// TIA Portal project "Canarias Skills" (V17) (continued)
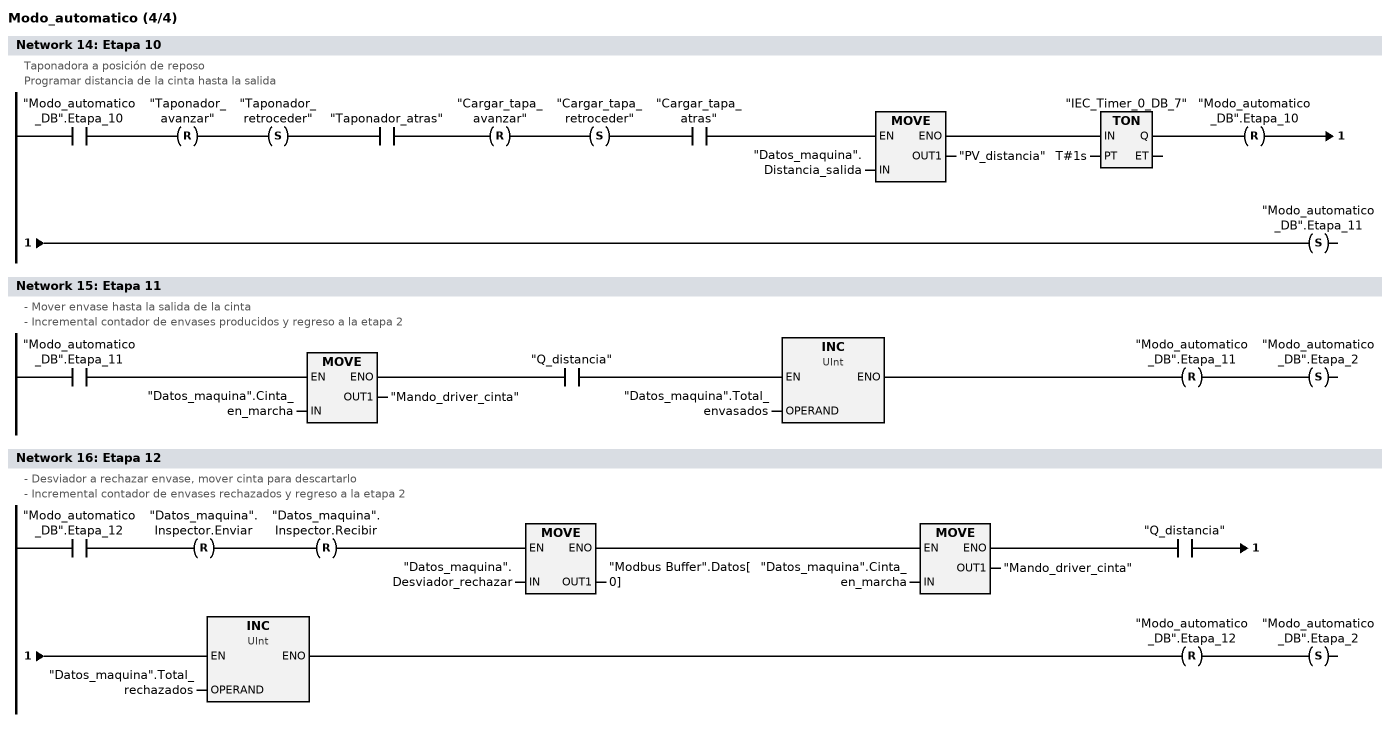
   IF "Modo_automatico_DB".Etapa_10 THEN
       "Taponador_avanzar" := FALSE;
       "Taponador_retroceder" := TRUE;
   END_IF;
   #_w1 := "Modo_automatico_DB".Etapa_10 AND "Taponador_atras";
   IF #_w1 THEN
       "Cargar_tapa_avanzar" := FALSE;
       "Cargar_tapa_retroceder" := TRUE;
   END_IF;
   #_w2 := #_w1 AND "Cargar_tapa_atras";
   IF #_w2 THEN "PV_distancia" := "Datos_maquina".Distancia_salida; END_IF;
   "IEC_Timer_0_DB_7".TON(IN := #_w2, PT := T#1s);
   IF "IEC_Timer_0_DB_7".Q THEN
       "Modo_automatico_DB".Etapa_10 := FALSE;
       "Modo_automatico_DB".Etapa_11 := TRUE;
   END_IF;
END_REGION

REGION Network 15: Etapa 11
   // - Mover envase hasta la salida de la cinta
   // - Incremental contador de envases producidos y regreso a la etapa 2
   RUNG wire#powerrail
      Contact( "Modo_automatico_DB".Etapa_11 )
      Move(in := "Datos_maquina".Cinta_en_marcha, out1 => "Mando_driver_cinta")
      Contact( "Q_distancia" )
      { S7_Templates := "DestType := UInt" } Inc( "Datos_maquina".Total_envasados )
      R_Coil( "Modo_automatico_DB".Etapa_11 )
      S_Coil( "Modo_automatico_DB".Etapa_2 )
   END_RUNG
   // the same network as SCL:
   IF "Modo_automatico_DB".Etapa_11 THEN "Mando_driver_cinta" := "Datos_maquina".Cinta_en_marcha; END_IF;
   IF "Modo_automatico_DB".Etapa_11 AND "Q_distancia" THEN
       "Datos_maquina".Total_envasados := "Datos_maquina".Total_envasados + 1;
   END_IF;
   #_w1 := "Modo_automatico_DB".Etapa_11 AND "Q_distancia";
   IF #_w1 THEN
       "Modo_automatico_DB".Etapa_11 := FALSE;
       "Modo_automatico_DB".Etapa_2 := TRUE;
   END_IF;
END_REGION

REGION Network 16: Etapa 12
   // - Desviador a rechazar envase, mover cinta para descartarlo
   // - Incremental contador de envases rechazados y regreso a la etapa 2
   RUNG wire#powerrail
      Contact( "Modo_automatico_DB".Etapa_12 )
      R_Coil( "Datos_maquina".Inspector.Enviar )
      R_Coil( "Datos_maquina".Inspector.Recibir )
      Move(in := "Datos_maquina".Desviador_rechazar, out1 => "Modbus Buffer".Datos[0])
      Move(in := "Datos_maquina".Cinta_en_marcha, out1 => "Mando_driver_cinta")
      Contact( "Q_distancia" )
      { S7_Templates := "DestType := UInt" } Inc( "Datos_maquina".Total_rechazados )
      R_Coil( "Modo_automatico_DB".Etapa_12 )
      S_Coil( "Modo_automatico_DB".Etapa_2 )
   END_RUNG
   // the same network as SCL:
   IF "Modo_automatico_DB".Etapa_12 THEN
       "Datos_maquina".Inspector.Enviar := FALSE;
       "Datos_maquina".Inspector.Recibir := FALSE;
       "Modbus Buffer".Datos[0] := "Datos_maquina".Desviador_rechazar;
       "Mando_driver_cinta" := "Datos_maquina".Cinta_en_marcha;
   END_IF;
   IF "Modo_automatico_DB".Etapa_12 AND "Q_distancia" THEN
       "Datos_maquina".Total_rechazados := "Datos_maquina".Total_rechazados + 1;
   END_IF;
   #_w1 := "Modo_automatico_DB".Etapa_12 AND "Q_distancia";
   IF #_w1 THEN
       "Modo_automatico_DB".Etapa_12 := FALSE;
       "Modo_automatico_DB".Etapa_2 := TRUE;
   END_IF;
END_REGION
END_FUNCTION_BLOCK

FUNCTION "Inicializar maquina" : Void   // FC1, LAD
{ S7_Optimized_Access := 'TRUE' }
VERSION : 0.1
BEGIN

REGION Network 1
   // Variador cinta, en servicio y detenido
   // Desviador en posición de aceptar envase
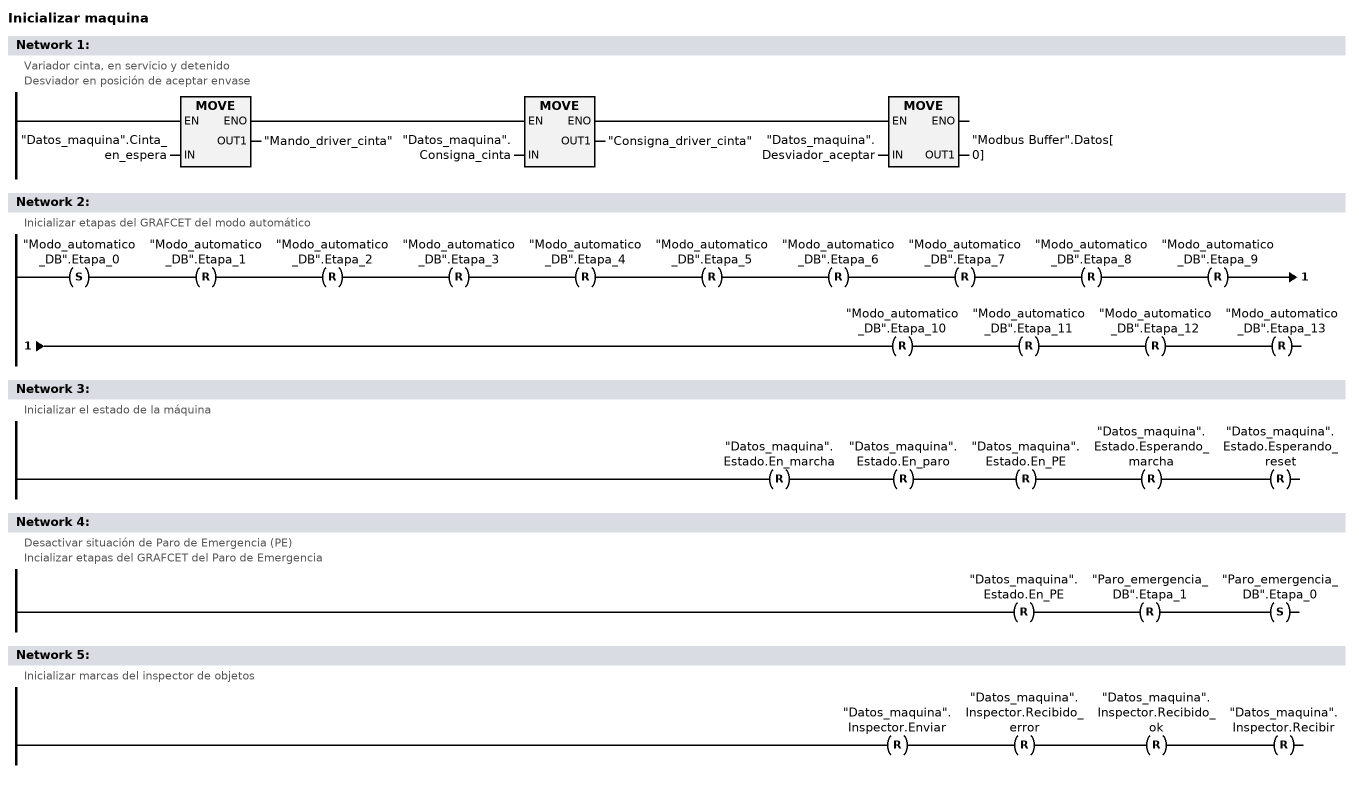
   RUNG wire#powerrail
      Move(in := "Datos_maquina".Cinta_en_espera, out1 => "Mando_driver_cinta")
      Move(in := "Datos_maquina".Consigna_cinta, out1 => "Consigna_driver_cinta")
      Move(in := "Datos_maquina".Desviador_aceptar, out1 => "Modbus Buffer".Datos[0])
   END_RUNG
   // the same network as SCL:
   "Mando_driver_cinta" := "Datos_maquina".Cinta_en_espera;
   "Consigna_driver_cinta" := "Datos_maquina".Consigna_cinta;
   "Modbus Buffer".Datos[0] := "Datos_maquina".Desviador_aceptar;
END_REGION

REGION Network 2
   // Inicializar etapas del GRAFCET del modo automático
   RUNG wire#powerrail
      S_Coil( "Modo_automatico_DB".Etapa_0 )
      R_Coil( "Modo_automatico_DB".Etapa_1 )
      R_Coil( "Modo_automatico_DB".Etapa_2 )
      R_Coil( "Modo_automatico_DB".Etapa_3 )
      R_Coil( "Modo_automatico_DB".Etapa_4 )
      R_Coil( "Modo_automatico_DB".Etapa_5 )
      R_Coil( "Modo_automatico_DB".Etapa_6 )
      R_Coil( "Modo_automatico_DB".Etapa_7 )
      R_Coil( "Modo_automatico_DB".Etapa_8 )
      R_Coil( "Modo_automatico_DB".Etapa_9 )
      R_Coil( "Modo_automatico_DB".Etapa_10 )
      R_Coil( "Modo_automatico_DB".Etapa_11 )
      R_Coil( "Modo_automatico_DB".Etapa_12 )
      R_Coil( "Modo_automatico_DB".Etapa_13 )
   END_RUNG
   // the same network as SCL:
   "Modo_automatico_DB".Etapa_0 := TRUE;
   "Modo_automatico_DB".Etapa_1 := FALSE;
   "Modo_automatico_DB".Etapa_2 := FALSE;
   "Modo_automatico_DB".Etapa_3 := FALSE;
   "Modo_automatico_DB".Etapa_4 := FALSE;
   "Modo_automatico_DB".Etapa_5 := FALSE;
   "Modo_automatico_DB".Etapa_6 := FALSE;
   "Modo_automatico_DB".Etapa_7 := FALSE;
   "Modo_automatico_DB".Etapa_8 := FALSE;
   "Modo_automatico_DB".Etapa_9 := FALSE;
   "Modo_automatico_DB".Etapa_10 := FALSE;
   "Modo_automatico_DB".Etapa_11 := FALSE;
   "Modo_automatico_DB".Etapa_12 := FALSE;
   "Modo_automatico_DB".Etapa_13 := FALSE;
END_REGION

REGION Network 3
   // Inicializar el estado de la máquina
   RUNG wire#powerrail
      R_Coil( "Datos_maquina".Estado.En_marcha )
      R_Coil( "Datos_maquina".Estado.En_paro )
      R_Coil( "Datos_maquina".Estado.En_PE )
      R_Coil( "Datos_maquina".Estado.Esperando_marcha )
      R_Coil( "Datos_maquina".Estado.Esperando_reset )
   END_RUNG
   // the same network as SCL:
   "Datos_maquina".Estado.En_marcha := FALSE;
   "Datos_maquina".Estado.En_paro := FALSE;
   "Datos_maquina".Estado.En_PE := FALSE;
   "Datos_maquina".Estado.Esperando_marcha := FALSE;
   "Datos_maquina".Estado.Esperando_reset := FALSE;
END_REGION

REGION Network 4
   // Desactivar situación de Paro de Emergencia (PE)
   // Incializar etapas del GRAFCET del Paro de Emergencia
   RUNG wire#powerrail
      R_Coil( "Datos_maquina".Estado.En_PE )
      R_Coil( "Paro_emergencia_DB".Etapa_1 )
      S_Coil( "Paro_emergencia_DB".Etapa_0 )
   END_RUNG
   // the same network as SCL:
   "Datos_maquina".Estado.En_PE := FALSE;
   "Paro_emergencia_DB".Etapa_1 := FALSE;
   "Paro_emergencia_DB".Etapa_0 := TRUE;
END_REGION

REGION Network 5
   // Inicializar marcas del inspector de objetos
   RUNG wire#powerrail
      R_Coil( "Datos_maquina".Inspector.Enviar )
      R_Coil( "Datos_maquina".Inspector.Recibido_error )
      R_Coil( "Datos_maquina".Inspector.Recibido_ok )
      R_Coil( "Datos_maquina".Inspector.Recibir )
   END_RUNG
   // the same network as SCL:
   "Datos_maquina".Inspector.Enviar := FALSE;
   "Datos_maquina".Inspector.Recibido_error := FALSE;
   "Datos_maquina".Inspector.Recibido_ok := FALSE;
   "Datos_maquina".Inspector.Recibir := FALSE;
END_REGION
END_FUNCTION

FUNCTION "Modo manual" : Void   // FC2, LAD
{ S7_Optimized_Access := 'TRUE' }
VERSION : 0.1
BEGIN

REGION Network 1: Maniobra manual de la neumática desde HMI
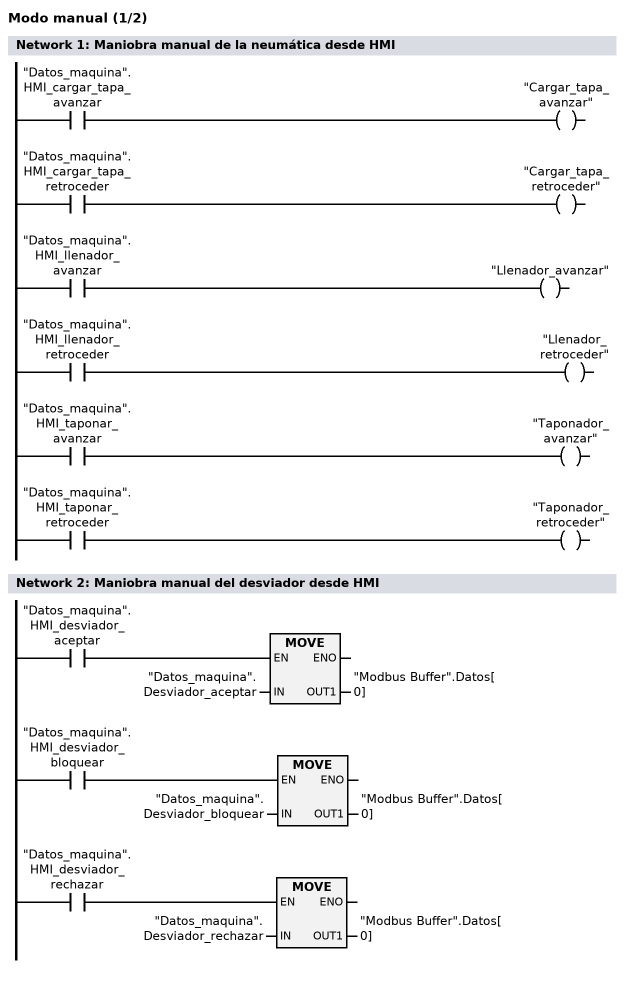
   RUNG wire#powerrail
      Contact( "Datos_maquina".HMI_cargar_tapa_avanzar )
      Coil( "Cargar_tapa_avanzar" )
   END_RUNG
   RUNG wire#powerrail
      Contact( "Datos_maquina".HMI_cargar_tapa_retroceder )
      Coil( "Cargar_tapa_retroceder" )
   END_RUNG
   RUNG wire#powerrail
      Contact( "Datos_maquina".HMI_llenador_avanzar )
      Coil( "Llenador_avanzar" )
   END_RUNG
   RUNG wire#powerrail
      Contact( "Datos_maquina".HMI_llenador_retroceder )
      Coil( "Llenador_retroceder" )
   END_RUNG
   RUNG wire#powerrail
      Contact( "Datos_maquina".HMI_taponar_avanzar )
      Coil( "Taponador_avanzar" )
   END_RUNG
   RUNG wire#powerrail
      Contact( "Datos_maquina".HMI_taponar_retroceder )
      Coil( "Taponador_retroceder" )
   END_RUNG
   // the same network as SCL:
   "Cargar_tapa_avanzar" := "Datos_maquina".HMI_cargar_tapa_avanzar;
   "Cargar_tapa_retroceder" := "Datos_maquina".HMI_cargar_tapa_retroceder;
   "Llenador_avanzar" := "Datos_maquina".HMI_llenador_avanzar;
   "Llenador_retroceder" := "Datos_maquina".HMI_llenador_retroceder;
   "Taponador_avanzar" := "Datos_maquina".HMI_taponar_avanzar;
   "Taponador_retroceder" := "Datos_maquina".HMI_taponar_retroceder;
END_REGION

REGION Network 2: Maniobra manual del desviador desde HMI
   RUNG wire#powerrail
      Contact( "Datos_maquina".HMI_desviador_aceptar )
      Move(in := "Datos_maquina".Desviador_aceptar, out1 => "Modbus Buffer".Datos[0])
   END_RUNG
   RUNG wire#powerrail
      Contact( "Datos_maquina".HMI_desviador_bloquear )
      Move(in := "Datos_maquina".Desviador_bloquear, out1 => "Modbus Buffer".Datos[0])
   END_RUNG
   RUNG wire#powerrail
      Contact( "Datos_maquina".HMI_desviador_rechazar )
      Move(in := "Datos_maquina".Desviador_rechazar, out1 => "Modbus Buffer".Datos[0])
   END_RUNG
   // the same network as SCL:
   IF "Datos_maquina".HMI_desviador_aceptar THEN
       "Modbus Buffer".Datos[0] := "Datos_maquina".Desviador_aceptar;
   END_IF;
   IF "Datos_maquina".HMI_desviador_bloquear THEN
       "Modbus Buffer".Datos[0] := "Datos_maquina".Desviador_bloquear;
   END_IF;
   IF "Datos_maquina".HMI_desviador_rechazar THEN
       "Modbus Buffer".Datos[0] := "Datos_maquina".Desviador_rechazar;
   END_IF;
END_REGION

REGION Network 3: Maniobras en modo manual del driver de la cinta
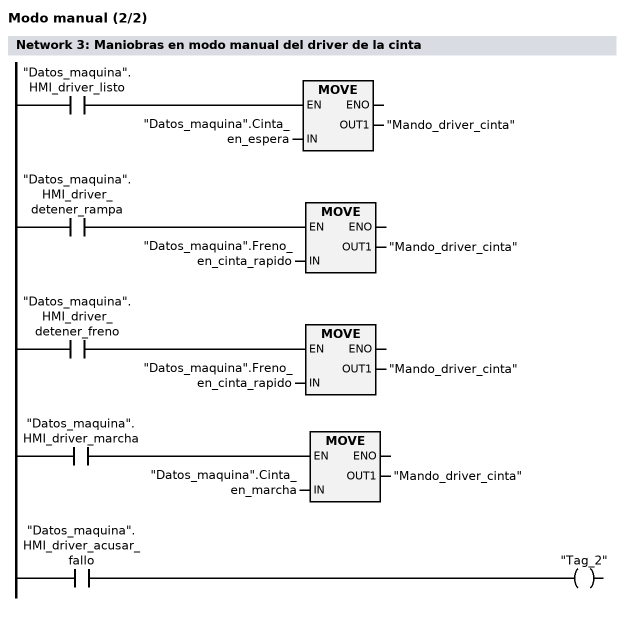
   RUNG wire#powerrail
      Contact( "Datos_maquina".HMI_driver_listo )
      Move(in := "Datos_maquina".Cinta_en_espera, out1 => "Mando_driver_cinta")
   END_RUNG
   RUNG wire#powerrail
      Contact( "Datos_maquina".HMI_driver_detener_rampa )
      Move(in := "Datos_maquina".Freno_en_cinta_rapido, out1 => "Mando_driver_cinta")
   END_RUNG
   RUNG wire#powerrail
      Contact( "Datos_maquina".HMI_driver_detener_freno )
      Move(in := "Datos_maquina".Freno_en_cinta_rapido, out1 => "Mando_driver_cinta")
   END_RUNG
   RUNG wire#powerrail
      Contact( "Datos_maquina".HMI_driver_marcha )
      Move(in := "Datos_maquina".Cinta_en_marcha, out1 => "Mando_driver_cinta")
   END_RUNG
   RUNG wire#powerrail
      Contact( "Datos_maquina".HMI_driver_acusar_fallo )
      Coil( "Tag_2" )
   END_RUNG
   // the same network as SCL:
   IF "Datos_maquina".HMI_driver_listo THEN "Mando_driver_cinta" := "Datos_maquina".Cinta_en_espera; END_IF;
   IF "Datos_maquina".HMI_driver_detener_rampa THEN
       "Mando_driver_cinta" := "Datos_maquina".Freno_en_cinta_rapido;
   END_IF;
   IF "Datos_maquina".HMI_driver_detener_freno THEN
       "Mando_driver_cinta" := "Datos_maquina".Freno_en_cinta_rapido;
   END_IF;
   IF "Datos_maquina".HMI_driver_marcha THEN "Mando_driver_cinta" := "Datos_maquina".Cinta_en_marcha; END_IF;
   "Tag_2" := "Datos_maquina".HMI_driver_acusar_fallo;
END_REGION
END_FUNCTION

FUNCTION "Actualizar alarmas" : Void   // FC3, LAD
{ S7_Optimized_Access := 'TRUE' }
VERSION : 0.1
BEGIN

REGION Network 1
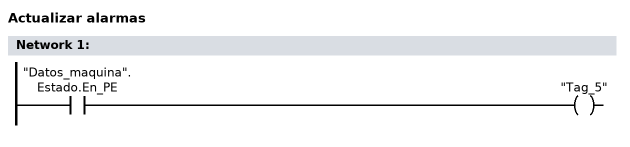
   RUNG wire#powerrail
      Contact( "Datos_maquina".Estado.En_PE )
      Coil( "Tag_5" )
   END_RUNG
   // the same network as SCL:
   "Tag_5" := "Datos_maquina".Estado.En_PE;
END_REGION
END_FUNCTION

ORGANIZATION_BLOCK "Main"   // OB1, LAD, ProgramCycle
TITLE = "Main Program Sweep (Cycle)"
{ S7_Optimized_Access := 'TRUE' }
VERSION : 0.1
   VAR_INPUT
      Initial_Call : Bool;   // Initial call of this OB
      Remanence : Bool;   // =True, if remanent data are available
   END_VAR
   VAR_TEMP
      aux : Int;
   END_VAR
BEGIN

REGION Network 1: Desviador de envases
   // Arduino UNO Modbus TCP, controla el servo del desviador de envases.
   // La posición del desviador se ajusta en DB3.DW0 "Modbus Buffer".Datos[0]
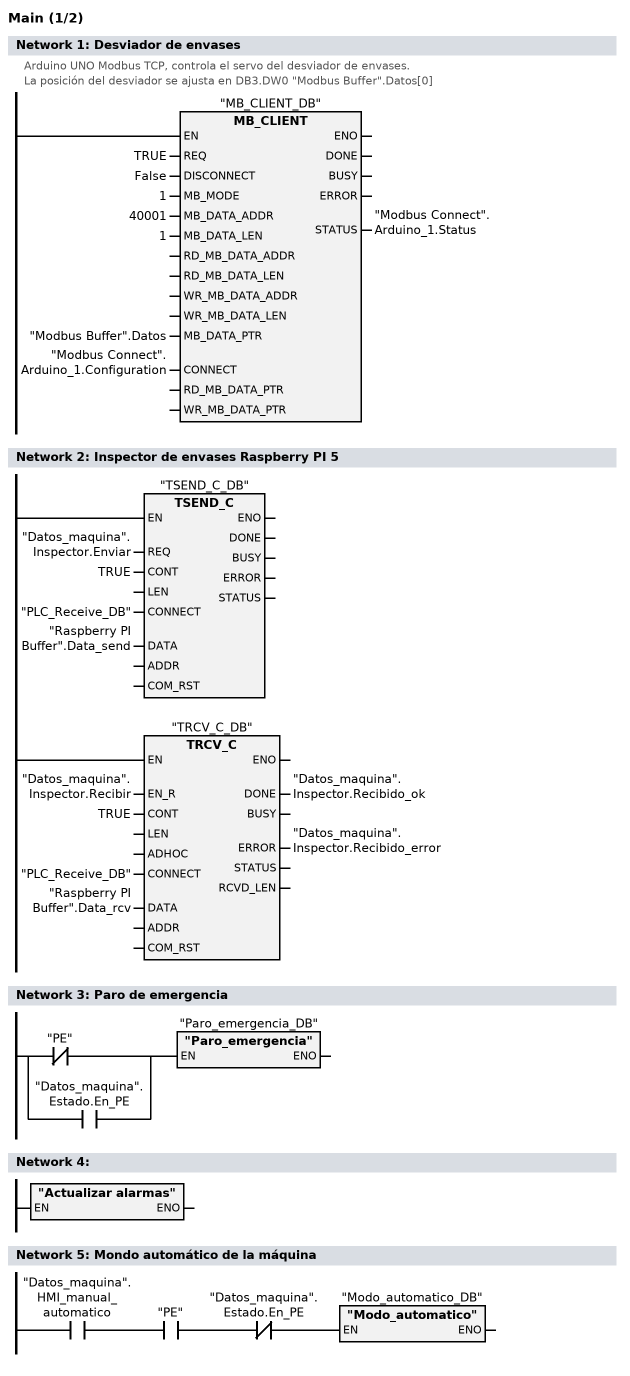
   "MB_CLIENT_DB"(REQ := TRUE,   // MB_CLIENT
                  DISCONNECT := False,
                  MB_MODE := 1,
                  MB_DATA_ADDR := 40001,
                  MB_DATA_LEN := 1,
                  MB_DATA_PTR := "Modbus Buffer".Datos,
                  CONNECT := "Modbus Connect".Arduino_1.Configuration,
                  STATUS => "Modbus Connect".Arduino_1.Status);
END_REGION

REGION Network 2: Inspector de envases Raspberry PI 5
   "TSEND_C_DB"(REQ := "Datos_maquina".Inspector.Enviar,   // TSEND_C
                CONT := TRUE,
                CONNECT := "PLC_Receive_DB",
                DATA := "Raspberry PI Buffer".Data_send);
   "TRCV_C_DB"(EN_R := "Datos_maquina".Inspector.Recibir,   // TRCV_C
               CONT := TRUE,
               CONNECT := "PLC_Receive_DB",
               DATA := "Raspberry PI Buffer".Data_rcv,
               DONE => "Datos_maquina".Inspector.Recibido_ok,
               ERROR => "Datos_maquina".Inspector.Recibido_error);
END_REGION

REGION Network 3: Paro de emergencia
   RUNG wire#powerrail
      I_Contact( "PE" )
      wire#w1
      "Paro_emergencia_DB"()
   END_RUNG
   RUNG wire#powerrail
      Contact( "Datos_maquina".Estado.En_PE )
   END_RUNG wire#w1
   // the same network as SCL:
   IF NOT "PE" OR "Datos_maquina".Estado.En_PE THEN
       "Paro_emergencia_DB"();   // "Paro_emergencia"
   END_IF;
END_REGION

REGION Network 4
   RUNG wire#powerrail
      "Actualizar alarmas"()
   END_RUNG
   // the same network as SCL:
   "Actualizar alarmas"();
END_REGION

REGION Network 5: Mondo automático de la máquina
   RUNG wire#powerrail
      Contact( "Datos_maquina".HMI_manual_automatico )
      Contact( "PE" )
      I_Contact( "Datos_maquina".Estado.En_PE )
      "Modo_automatico_DB"()
   END_RUNG
   // the same network as SCL:
   IF "Datos_maquina".HMI_manual_automatico AND "PE" AND NOT "Datos_maquina".Estado.En_PE THEN
       "Modo_automatico_DB"();   // "Modo_automatico"
   END_IF;
END_REGION

REGION Network 6: Modo manual de la máquina
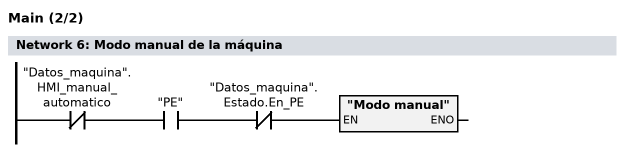
   RUNG wire#powerrail
      I_Contact( "Datos_maquina".HMI_manual_automatico )
      Contact( "PE" )
      I_Contact( "Datos_maquina".Estado.En_PE )
      "Modo manual"()
   END_RUNG
   // the same network as SCL:
   IF NOT "Datos_maquina".HMI_manual_automatico AND "PE" AND NOT "Datos_maquina".Estado.En_PE THEN
       "Modo manual"();
   END_IF;
END_REGION
END_ORGANIZATION_BLOCK

ORGANIZATION_BLOCK "Startup"   // OB100, LAD, Startup
TITLE = "Complete Restart"
{ S7_Optimized_Access := 'TRUE' }
VERSION : 0.1
   VAR_INPUT
      LostRetentive : Bool;   // True if retentive data are lost
      LostRTC : Bool;   // True if date and time are lost
   END_VAR
   VAR_TEMP   // added for the SCL form of the ladder/FBD networks
      _w1 : Bool;
   END_VAR
BEGIN

REGION Network 1: Marcha desde el HMI
   // Desactivar Marcha, Paro y Reset del HMI
   // Activar modo automatico del HMI
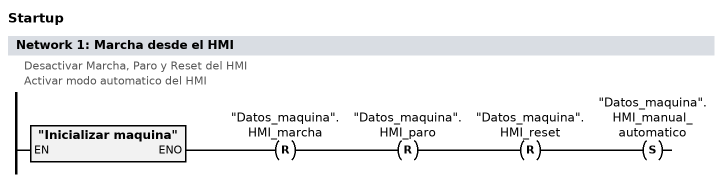
   RUNG wire#powerrail
      "Inicializar maquina"()
      R_Coil( "Datos_maquina".HMI_marcha )
      R_Coil( "Datos_maquina".HMI_paro )
      R_Coil( "Datos_maquina".HMI_reset )
      S_Coil( "Datos_maquina".HMI_manual_automatico )
   END_RUNG
   // the same network as SCL:
   "Inicializar maquina"(ENO => #_w1);
   IF #_w1 THEN
       "Datos_maquina".HMI_marcha := FALSE;
       "Datos_maquina".HMI_paro := FALSE;
       "Datos_maquina".HMI_reset := FALSE;
       "Datos_maquina".HMI_manual_automatico := TRUE;
   END_IF;
END_REGION
END_ORGANIZATION_BLOCK

(* ===== HMI "HMI_RT_1" =====
system functions are stored by id; their names below are inferred from use
connection "HMI_Connection_1": ETHERNET, SMART_S7_1200_OMS

HMI tags "Default tag table"
   "Tag_ScreenNumber" : UInt, internal
   "Datos_maquina_HMI_llenador_avanzar" : Bool = PLC Datos_maquina.HMI_llenador_avanzar, 1 s
   "Datos_maquina_HMI_llenador_retroceder" : Bool = PLC Datos_maquina.HMI_llenador_retroceder, 1 s
   "Datos_maquina_HMI_cargar_tapa_avanzar" : Bool = PLC Datos_maquina.HMI_cargar_tapa_avanzar, 1 s
   "Datos_maquina_HMI_cargar_tapa_retroceder" : Bool = PLC Datos_maquina.HMI_cargar_tapa_retroceder, 1 s
   "Datos_maquina_HMI_taponar_avanzar" : Bool = PLC Datos_maquina.HMI_taponar_avanzar, 1 s
   "Datos_maquina_HMI_taponar_retroceder" : Bool = PLC Datos_maquina.HMI_taponar_retroceder, 1 s
   "Datos_maquina_HMI_desviador_bloquear" : Bool = PLC Datos_maquina.HMI_desviador_bloquear, 1 s
   "Datos_maquina_HMI_desviador_rechazar" : Bool = PLC Datos_maquina.HMI_desviador_rechazar, 1 s
   "Datos_maquina_HMI_desviador_aceptar" : Bool = PLC Datos_maquina.HMI_desviador_aceptar, 1 s
   "Datos_maquina_HMI_driver_listo" : Bool = PLC Datos_maquina.HMI_driver_listo, 1 s
   "Datos_maquina_HMI_driver_marcha" : Bool = PLC Datos_maquina.HMI_driver_marcha, 1 s
   "Datos_maquina_HMI_driver_detener_rampa" : Bool = PLC Datos_maquina.HMI_driver_detener_rampa, 1 s
   "Datos_maquina_HMI_driver_detener_freno" : Bool = PLC Datos_maquina.HMI_driver_detener_freno, 1 s
   "Datos_maquina_HMI_driver_acusar_fallo" : Bool = PLC Datos_maquina.HMI_driver_acusar_fallo, 1 s
   "Datos_maquina_Total_envasados" : Word = PLC Datos_maquina.Total_envasados, 1 s
   "Datos_maquina_Total_rechazados" : Word = PLC Datos_maquina.Total_rechazados, 1 s
   "Datos_maquina_Distancia_inspeccion" : Word = PLC Datos_maquina.Distancia_inspeccion, 1 s
   "Datos_maquina_Distancia_desviador" : Word = PLC Datos_maquina.Distancia_desviador, 1 s
   "Datos_maquina_Distancia_llenadora" : Word = PLC Datos_maquina.Distancia_llenadora, 1 s
   "Datos_maquina_Distancia_taponadora" : Word = PLC Datos_maquina.Distancia_taponadora, 1 s
   "Datos_maquina_Distancia_salida" : Word = PLC Datos_maquina.Distancia_salida, 1 s
   "Datos_maquina_HMI_manual_automatico" : Bool = PLC Datos_maquina.HMI_manual_automatico, 1 s
   "Datos_maquina_HMI_marcha" : Bool = PLC Datos_maquina.HMI_marcha, 1 s
   "Datos_maquina_HMI_paro" : Bool = PLC Datos_maquina.HMI_paro, 1 s
   "Datos_maquina_HMI_reset" : Bool = PLC Datos_maquina.HMI_reset, 1 s
   "Datos_maquina_Desviador_bloquear" : Word = PLC Datos_maquina.Desviador_bloquear, 1 s
   "Datos_maquina_Desviador_aceptar" : Word = PLC Datos_maquina.Desviador_aceptar, 1 s
   "Datos_maquina_Desviador_rechazar" : Word = PLC Datos_maquina.Desviador_rechazar, 1 s
   "PV_distancia" : Word = PLC PV_distancia AT %MW212, 1 s
   "CV_distancia" : Word = PLC CV_distancia AT %MW214, 1 s
   "Datos_maquina_Estado_Esperando_marcha" : Bool = PLC Datos_maquina.Estado.Esperando_marcha, 1 s
   "Datos_maquina_Estado_En_paro" : Bool = PLC Datos_maquina.Estado.En_paro, 1 s
   "Datos_maquina_Estado_Esperando_reset" : Bool = PLC Datos_maquina.Estado.Esperando_reset, 1 s
   "Alarmas" : Word = PLC Alarmas AT %MW100, 1 s
   "ACK_alarmas" : Word = PLC ACK_alarmas AT %MW102, 1 s

discrete alarms
   1: 'Parada de emergencia', class Errors, trigger "Alarmas" bit 8

Template "Template_1" 800x480
   Button "Exit" at 714,429 size 71x50; TextOff 'Exit'; PictureOff "ExitRuntime_KTP700_Basic_PN_TR"; PictureOn "ExitRuntime_KTP700_Basic_PN_TR"
      on Release: StopRuntime(0)
   Button "Template_Button" at 614,429 size 71x50; TextOff 'Text'
   Button "Template_Button_1" at 514,429 size 71x50; TextOff 'Text'
   Button "Template_Button_2" at 414,429 size 71x50; TextOff 'Text'
   Button "Template_Button_3" at 314,429 size 71x50; TextOff 'Text'
   Button "Log on" at 214,429 size 71x50; TextOff 'Log on'; PictureOff "Login_KTP700_Basic_PN_TR"; PictureOn "Login_KTP700_Basic_PN_TR"
      on Release: function_a2a04561()
   Button "Alarms" at 114,429 size 71x50; TextOff 'Alarms'; PictureOff "AlarmDisplay_KTP700_Basic_PN_TR"; PictureOn "AlarmDisplay_KTP700_Basic_PN_TR"
      on Release: function_ef3f5d25("Alarm window_Unacknowledged", -1)
   Button "Start screen" at 14,429 size 71x50; TextOff 'Start screen'; PictureOff "NavigateHome_KTP700_Basic_PN_TR"; PictureOn "NavigateHome_KTP700_Basic_PN_TR"
      on Release: ActivateScreen("Inicio", 0)
   SymbolicIOField "Symbolic_IO_Field_Screen" at 170,9 size 523x33; TextOff '0'; TextOn '1'; TextList "TextList_ScreenNames"
      ProcessValue <- "Tag_ScreenNumber"
      on Change: ActivateScreenByNumber("Tag_ScreenNumber", 0)
   DateTimeField "HmiScreenItemData" at 695,25 size 105x25
   DateTimeField "HmiScreenItemData_1" at 695,0 size 105x25
   GraphicView "Logo" at 0,0 size 168x51; Picture "Logo of HMI_1"
   AlarmView "Template_Alarm view_1" at 156,74 size 623x300

screen "Inicio" 800x480, template "Template_1"
   on GenerateScreen: SetTag("Tag_ScreenNumber", 1)
   TextField "HmiScreenItemData_4" at 146,240 size 640x40; Text 'Envasadora de productos cosméticos'
   Button "HmiScreenItemData" at 36,87 size 159x47; TextOff 'Modo Manual'; PictureOff "Navigates to Modo Manual for KTP700 Basic+ PN 17.0.0.0"; PictureOn "Navigates to Modo Manual for KTP700 Basic+ PN 17.0.0.0"; Authorization "Maniobrar"
      on Release: ActivateScreen("Modo Manual", 0)
      Visibility <- "Datos_maquina_HMI_manual_automatico"
   Button "HmiScreenItemData_1" at 36,146 size 159x47; TextOff 'Modo Automático'; PictureOff "Navigates to Modo Automático for KTP700 Basic+ PN 17.0.0.0"; PictureOn "Navigates to Modo Automático for KTP700 Basic+ PN 17.0.0.0"; Authorization "Maniobrar"
      on Release: ActivateScreen("Modo Automático", 0)
   Button "HmiScreenItemData_2" at 36,205 size 159x47; TextOff 'Configuración máquina'; PictureOff "Navigates to Configuración máquina for KTP700 Basic+ PN 17.0.0.0"; PictureOn "Navigates to Configuración máquina for KTP700 Basic+ PN 17.0.0.0"; Authorization "Configurar"
      on Release: ActivateScreen("Configuración máquina", 0)
      Visibility <- "Datos_maquina_HMI_manual_automatico"
   Button "HmiScreenItemData_3" at 36,264 size 159x47; TextOff 'Estadísticas'; PictureOff "Navigates to Estadísticas for KTP700 Basic+ PN 17.0.0.0"; PictureOn "Navigates to Estadísticas for KTP700 Basic+ PN 17.0.0.0"; Authorization "Observar"
      on Release: ActivateScreen("Estadísticas", 0)
   Button "HmiScreenItemData_5" at 36,323 size 159x47; TextOff 'Sistema'; PictureOff "Navigates to System screens for KTP700 Basic+ PN 17.0.0.0"; PictureOn "Navigates to System screens for KTP700 Basic+ PN 17.0.0.0"; Authorization "Configurar"
      on Release: ActivateScreen("Sistema", 0)
   TextField "HmiScreenItemData_6" at 145,279 size 640x25; Text 'Canarias Skills 2024'
   GraphicView "Graphic view_1" at 216,87 size 510x137; Picture "Logo centro"

screen "Modo Manual" 800x480, template "Template_1"
   on GenerateScreen: SetTag("Tag_ScreenNumber", 2)
   Button "Back" at 15,355 size 150x45; TextOff 'Inicio'; TextOn 'Back'
      on Release: ActivateScreen("Inicio", 0)
   Button "Button_1" at 183,83 size 170x45; TextOff 'Llenador +'
      on Press: SetBit("Datos_maquina_HMI_llenador_avanzar")
      on Release: ResetBit("Datos_maquina_HMI_llenador_avanzar")
   Button "Button_2" at 183,136 size 170x45; TextOff 'Llenador -'
      on Release: ResetBit("Datos_maquina_HMI_llenador_retroceder")
      on Press: SetBit("Datos_maquina_HMI_llenador_retroceder")
   Button "Button_3" at 183,193 size 170x45; TextOff 'Sacar tapa +'
      on Release: ResetBit("Datos_maquina_HMI_cargar_tapa_avanzar")
      on Press: SetBit("Datos_maquina_HMI_cargar_tapa_avanzar")
   Button "Button_4" at 183,246 size 170x45; TextOff 'Sacar tapa -'
      on Release: ResetBit("Datos_maquina_HMI_cargar_tapa_retroceder")
      on Press: SetBit("Datos_maquina_HMI_cargar_tapa_retroceder")
   Button "Button_5" at 183,302 size 170x45; TextOff 'Taponador +'
      on Release: ResetBit("Datos_maquina_HMI_taponar_avanzar")
      on Press: SetBit("Datos_maquina_HMI_taponar_avanzar")
   Button "Button_6" at 183,355 size 170x45; TextOff 'Taponador -'
      on Release: ResetBit("Datos_maquina_HMI_taponar_retroceder")
      on Press: SetBit("Datos_maquina_HMI_taponar_retroceder")
   Button "Button_7" at 374,136 size 170x45; TextOff 'Desviador bloquear'
      on Press: SetBit("Datos_maquina_HMI_desviador_bloquear")
      on Release: ResetBit("Datos_maquina_HMI_desviador_bloquear")
   Button "Button_8" at 374,193 size 170x45; TextOff 'Desviador descartar'
      on Release: ResetBit("Datos_maquina_HMI_desviador_rechazar")
      on Press: SetBit("Datos_maquina_HMI_desviador_rechazar")
   Button "Button_9" at 374,246 size 170x45; TextOff 'Desviador aceptar'
      on Release: ResetBit("Datos_maquina_HMI_desviador_aceptar")
      on Press: SetBit("Datos_maquina_HMI_desviador_aceptar")
   Button "Button_10" at 564,136 size 170x45; TextOff 'Cinta preparada'
      on Release: ResetBit("Datos_maquina_HMI_driver_listo")
      on Press: SetBit("Datos_maquina_HMI_driver_listo")
   Button "Button_11" at 564,193 size 170x45; TextOff 'Marcha cinta'
      on Release: ResetBit("Datos_maquina_HMI_driver_marcha")
      on Press: SetBit("Datos_maquina_HMI_driver_marcha")
   Button "Button_12" at 564,246 size 170x45; TextOff 'Parar por rampa'
      on Release: ResetBit("Datos_maquina_HMI_driver_detener_rampa")
      on Press: SetBit("Datos_maquina_HMI_driver_detener_rampa")
   Button "Button_13" at 564,302 size 170x45; TextOff 'Parar por freno'
      on Release: ResetBit("Datos_maquina_HMI_driver_detener_freno")
      on Press: SetBit("Datos_maquina_HMI_driver_detener_freno")
   Button "Button_14" at 564,355 size 170x45; TextOff 'Acusar fallo cinta'
      on Release: ResetBit("Datos_maquina_HMI_driver_acusar_fallo")
      on Press: SetBit("Datos_maquina_HMI_driver_acusar_fallo")

screen "Modo Automático" 800x480, template "Template_1"
   on GenerateScreen: SetTag("Tag_ScreenNumber", 3)
   Button "Back" at 12,353 size 165x50; TextOff 'Inicio'; TextOn 'Back'
      on Release: ActivateScreen("Inicio", 0)
   Switch "Switch_1" at 12,90 size 165x50; CaptionText 'Switch'; TextOff 'Manual'; TextOn 'Auto'
      on SwitchOn: SetBit("Datos_maquina_HMI_manual_automatico")
      on SwitchOff: ResetBit("Datos_maquina_HMI_manual_automatico")
      ProcessValue <- "Datos_maquina_HMI_manual_automatico"
   Button "Button_1" at 13,146 size 165x50; TextOff 'Marcha'
      on Press: SetBit("Datos_maquina_HMI_marcha")
      on Release: ResetBit("Datos_maquina_HMI_marcha")
      Visibility <- "Datos_maquina_HMI_manual_automatico"
      Appearance <- "Datos_maquina_Estado_Esperando_marcha"
   Button "Button_2" at 13,201 size 165x50; TextOff 'Paro'
      on Press: SetBit("Datos_maquina_HMI_paro")
      on Release: ResetBit("Datos_maquina_HMI_paro")
      Visibility <- "Datos_maquina_HMI_manual_automatico"
      Appearance <- "Datos_maquina_Estado_En_paro"
   Button "Button_3" at 13,257 size 165x50; TextOff 'Reset'
      on Press: SetBit("Datos_maquina_HMI_reset")
      on Release: ResetBit("Datos_maquina_HMI_reset")
      Appearance <- "Datos_maquina_Estado_Esperando_reset"
   IOField "I/O field_1" at 313,178 size 96x32; FormatPattern 99999
      ProcessValue <- "Datos_maquina_Total_envasados"
   IOField "I/O field_2" at 313,233 size 96x32; FormatPattern 99999
      ProcessValue <- "Datos_maquina_Total_rechazados"
   TextField "Text field_1" at 311,156 size 138x23; Text 'Total envasados'
   TextField "Text field_2" at 311,212 size 145x23; Text 'Total rechazados'
   IOField "I/O field_3" at 564,180 size 96x32; FormatPattern 99999
      ProcessValue <- "PV_distancia"
   TextField "Text field_3" at 561,160 size 105x23; Text 'PV distancia'
   IOField "I/O field_4" at 564,235 size 96x32; FormatPattern 99999
      ProcessValue <- "CV_distancia"
   TextField "Text field_4" at 561,215 size 125x23; Text 'Contador cinta'

screen "Configuración máquina" 800x480, template "Template_1"
   on GenerateScreen: SetTag("Tag_ScreenNumber", 4)
   TextField "HmiScreenItemData" at 78,53 size 640x25; Text 'Configuración máquina'
   Button "Back" at 15,369 size 170x47; TextOff 'Inicio'; TextOn 'Back'
      on Release: ActivateScreen("Inicio", 0)
   IOField "I/O field_1" at 285,109 size 96x32; FormatPattern 99999
      ProcessValue <- "Datos_maquina_Distancia_inspeccion"
   IOField "I/O field_2" at 285,157 size 96x32; FormatPattern 99999
      ProcessValue <- "Datos_maquina_Distancia_desviador"
   IOField "I/O field_3" at 285,206 size 96x32; FormatPattern 99999
      ProcessValue <- "Datos_maquina_Distancia_llenadora"
   IOField "I/O field_4" at 285,254 size 96x32; FormatPattern 99999
      ProcessValue <- "Datos_maquina_Distancia_taponadora"
   IOField "I/O field_5" at 285,297 size 96x32; FormatPattern 99999
      ProcessValue <- "Datos_maquina_Distancia_salida"
   TextField "Text field_1" at 71,111 size 209x24; Text 'Distancia inspector (mm)'
   TextField "Text field_2" at 67,159 size 213x23; Text 'Distancia desviador (mm)'
   TextField "Text field_3" at 69,210 size 211x23; Text 'Distancia llenadora (mm)'
   TextField "Text field_4" at 52,256 size 228x23; Text 'Distancia taponadora (mm)'
   TextField "Text field_5" at 53,301 size 227x23; Text 'Distancia salida cinta (mm)'
   IOField "I/O field_6" at 617,109 size 96x32; FormatPattern 99999
      ProcessValue <- "Datos_maquina_Desviador_bloquear"
   IOField "I/O field_7" at 617,157 size 96x32; FormatPattern 99999
      ProcessValue <- "Datos_maquina_Desviador_rechazar"
   IOField "I/O field_8" at 617,206 size 96x32; FormatPattern 99999
      ProcessValue <- "Datos_maquina_Desviador_aceptar"
   TextField "Text field_6" at 420,111 size 191x23; Text 'Desviador bloquear (º)'
   TextField "Text field_7" at 421,159 size 190x23; Text 'Desviador rechazar (º)'
   TextField "Text field_8" at 430,210 size 181x23; Text 'Desviador aceptar (º)'
   Button "Button_7" at 543,259 size 170x45; TextOff 'Desviador bloquear'
      on Release: ResetBit("Datos_maquina_HMI_desviador_bloquear")
      on Press: SetBit("Datos_maquina_HMI_desviador_bloquear")
   Button "Button_8" at 543,316 size 170x45; TextOff 'Desviador descartar'
      on Release: ResetBit("Datos_maquina_HMI_desviador_rechazar")
      on Press: SetBit("Datos_maquina_HMI_desviador_rechazar")
   Button "Button_9" at 543,371 size 170x45; TextOff 'Desviador aceptar'
      on Release: ResetBit("Datos_maquina_HMI_desviador_aceptar")
      on Press: SetBit("Datos_maquina_HMI_desviador_aceptar")

screen "Estadísticas" 800x480, template "Template_1"
   on GenerateScreen: SetTag("Tag_ScreenNumber", 5)
   TextField "HmiScreenItemData" at 75,49 size 640x25; Text 'Estadísticas'
   Button "Back" at 16,371 size 169x47; TextOff 'Inicio'; TextOn 'Back'
      on Release: ActivateScreen("Inicio", 0)
   IOField "I/O field_1" at 456,147 size 96x32; FormatPattern 99999
      ProcessValue <- "Datos_maquina_Total_envasados"
   IOField "I/O field_2" at 456,198 size 96x32; FormatPattern 99999
      ProcessValue <- "Datos_maquina_Total_rechazados"
   TextField "Text field_1" at 314,152 size 138x23; Text 'Total envasados'
   TextField "Text field_2" at 307,203 size 145x23; Text 'Total rechazados'
   Button "Button_1" at 352,248 size 200x56; TextOff 'Borrar contadores'; Authorization "Borrado General"
      on Click: SetTag("Datos_maquina_Total_envasados", 0); SetTag("Datos_maquina_Total_rechazados", 0)

screen "Sistema" 800x480, template "Template_1"
   on GenerateScreen: SetTag("Tag_ScreenNumber", 6)
   Button "Back" at 30,359 size 159x47; TextOff 'Inicio'; TextOn 'Back'
      on Release: ActivateScreen("Inicio", 0)
   Button "HmiScreenItemData" at 30,111 size 159x47; TextOff 'SIMATIC PLC system diagnos...'; PictureOff "Navigates to SIMATIC PLC system diagnostics for KTP700 Basic+ PN 17.0.0.0"; PictureOn "Navigates to SIMATIC PLC system diagnostics for KTP700 Basic+ PN 17.0.0.0"
      on Release: ActivateScreen("SIMATIC PLC diagnósticos de sistema", 0)
   Button "HmiScreenItemData_1" at 30,170 size 159x47; TextOff 'Project information'; PictureOff "Navigates to Project information for KTP700 Basic+ PN 17.0.0.0"; PictureOn "Navigates to Project information for KTP700 Basic+ PN 17.0.0.0"
      on Release: ActivateScreen("Información del proyecto", 0)
   Button "HmiScreenItemData_2" at 30,229 size 159x47; TextOff 'User administration'; PictureOff "Navigates to User administration for KTP700 Basic+ PN 17.0.0.0"; PictureOn "Navigates to User administration for KTP700 Basic+ PN 17.0.0.0"
      on Release: ActivateScreen("Administración de usuarios", 0)
   Button "HmiScreenItemData_3" at 30,288 size 159x47; TextOff 'System information'; PictureOff "Navigates to System information for KTP700 Basic+ PN 17.0.0.0"; PictureOn "Navigates to System information for KTP700 Basic+ PN 17.0.0.0"
      on Release: ActivateScreen("Información del sistema", 0)
   Button "HmiScreenItemData_4" at 201,111 size 159x47; TextOff 'Different jobs'; PictureOff "Navigates to Different jobs for KTP700 Basic+ PN 17.0.0.0"; PictureOn "Navigates to Different jobs for KTP700 Basic+ PN 17.0.0.0"
      on Release: ActivateScreen("Otras tareas", 0)

screen "SIMATIC PLC diagnósticos de sistema" 800x480, template "Template_1"
   on GenerateScreen: SetTag("Tag_ScreenNumber", 7)
   SysDiagControl "HmiScreenItemData" at 1,51 size 796x321
   Button "Back" at 16,377 size 169x47; TextOff 'Inicio'; TextOn 'Back'
      on Release: ActivateScreen("Sistema", 0)

screen "Información del proyecto" 800x480, template "Template_1"
   on GenerateScreen: SetTag("Tag_ScreenNumber", 8)
   TextField "HmiScreenItemData" at 35,102 size 171x28; Text 'Project name:'
   TextField "HmiScreenItemData_1" at 241,102 size 524x28; Text 'Canarias Skills 2024'
   TextField "HmiScreenItemData_2" at 35,132 size 171x28; Text 'Created on:'
   TextField "HmiScreenItemData_3" at 241,132 size 524x28; Text '12/9/2022 1:26:35 PM'
   TextField "HmiScreenItemData_4" at 35,162 size 171x28; Text 'Author:'
   TextField "HmiScreenItemData_5" at 241,162 size 524x28; Text 'Curso de Especialización en Ciberseguridad en'
   TextField "HmiScreenItemData_6" at 35,217 size 171x28; Text 'Description:'
   TextField "HmiScreenItemData_7" at 241,217 size 524x28; Text 'Máquina envasadora de productos cosméticos'
   Button "Back" at 17,361 size 168x47; TextOff 'Inicio'; TextOn 'Back'
      on Release: ActivateScreen("Sistema", 0)
   TextField "HmiScreenItemData_8" at 241,190 size 524x28; Text 'Tecnologías de Operación (OT)'

screen "Administración de usuarios" 800x480, template "Template_1"
   on GenerateScreen: SetTag("Tag_ScreenNumber", 9)
   UserView "HmiScreenItemData" at 1,54 size 796x321
   Button "Back" at 16,379 size 168x47; TextOff 'Inicio'; TextOn 'Back'
      on Release: ActivateScreen("Sistema", 0)

screen "Información del sistema" 800x480, template "Template_1"
   on GenerateScreen: SetTag("Tag_ScreenNumber", 10)
   Button "Back" at 17,372 size 169x47; TextOff 'Inicio'; TextOn 'Back'
      on Release: ActivateScreen("Sistema", 0)
   GraphicView "Graphic view_1" at 191,61 size 602x354; Picture "Estructura de la red"

screen "Otras tareas" 800x480, template "Template_1"
   on GenerateScreen: SetTag("Tag_ScreenNumber", 11)
   Button "Online" at 36,80 size 159x47; TextOff 'Online'
      on Release: function_bb44b551(0)
   Button "Offline" at 36,139 size 159x47; TextOff 'Offline'
      on Release: function_bb44b551(1)
   Button "Transfer" at 36,198 size 159x47; TextOff 'Cargar proyecto'; TextOn 'Transfer'; Authorization "Configurar"
      on Release: function_bb44b551(2)
   Button "Toggle language" at 36,257 size 159x47; TextOff 'Cambiar idioma'; TextOn 'Toggle language'; Authorization "Configurar"
      on Release: function_fb9197e8(-1)
   Button "Stop Runtime" at 207,80 size 159x47; TextOff 'Stop Runtime'; Authorization "Configurar"
      on Release: StopRuntime(0)
   Button "Back" at 38,366 size 159x47; TextOff 'Inicio'; TextOn 'Back'
      on Release: ActivateScreen("Sistema", 0)
*)